// TIA Portal project "FS-DS-09" (V16) (continued)
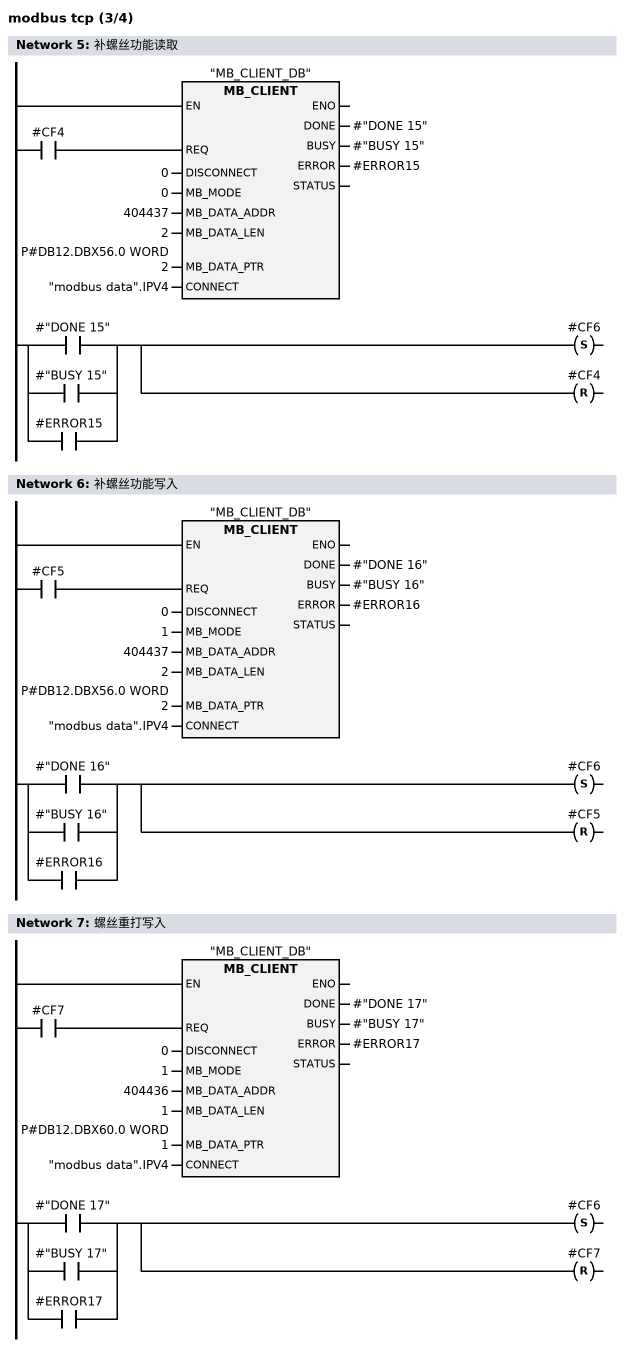
   "MB_CLIENT_DB"(REQ := #CF4,   // MB_CLIENT
                  DISCONNECT := 0,
                  MB_MODE := 0,
                  MB_DATA_ADDR := 404437,
                  MB_DATA_LEN := 2,
                  MB_DATA_PTR := P#DB12.DBX56.0 WORD 2,
                  CONNECT := "modbus data".IPV4,
                  DONE => #"DONE 15",
                  BUSY => #"BUSY 15",
                  ERROR => #ERROR15);
   IF #"DONE 15" OR #"BUSY 15" OR #ERROR15 THEN
       #CF6 := TRUE;
       #CF4 := FALSE;
   END_IF;
END_REGION

REGION Network 6: 补螺丝功能写入
   "MB_CLIENT_DB"(REQ := #CF5,   // MB_CLIENT
                  DISCONNECT := 0,
                  MB_MODE := 1,
                  MB_DATA_ADDR := 404437,
                  MB_DATA_LEN := 2,
                  MB_DATA_PTR := P#DB12.DBX56.0 WORD 2,
                  CONNECT := "modbus data".IPV4,
                  DONE => #"DONE 16",
                  BUSY => #"BUSY 16",
                  ERROR => #ERROR16);
   IF #"DONE 16" OR #"BUSY 16" OR #ERROR16 THEN
       #CF6 := TRUE;
       #CF5 := FALSE;
   END_IF;
END_REGION

REGION Network 7: 螺丝重打写入
   "MB_CLIENT_DB"(REQ := #CF7,   // MB_CLIENT
                  DISCONNECT := 0,
                  MB_MODE := 1,
                  MB_DATA_ADDR := 404436,
                  MB_DATA_LEN := 1,
                  MB_DATA_PTR := P#DB12.DBX60.0 WORD 1,
                  CONNECT := "modbus data".IPV4,
                  DONE => #"DONE 17",
                  BUSY => #"BUSY 17",
                  ERROR => #ERROR17);
   IF #"DONE 17" OR #"BUSY 17" OR #ERROR17 THEN
       #CF6 := TRUE;
       #CF7 := FALSE;
   END_IF;
END_REGION

REGION Network 8: 回原位标志位写入
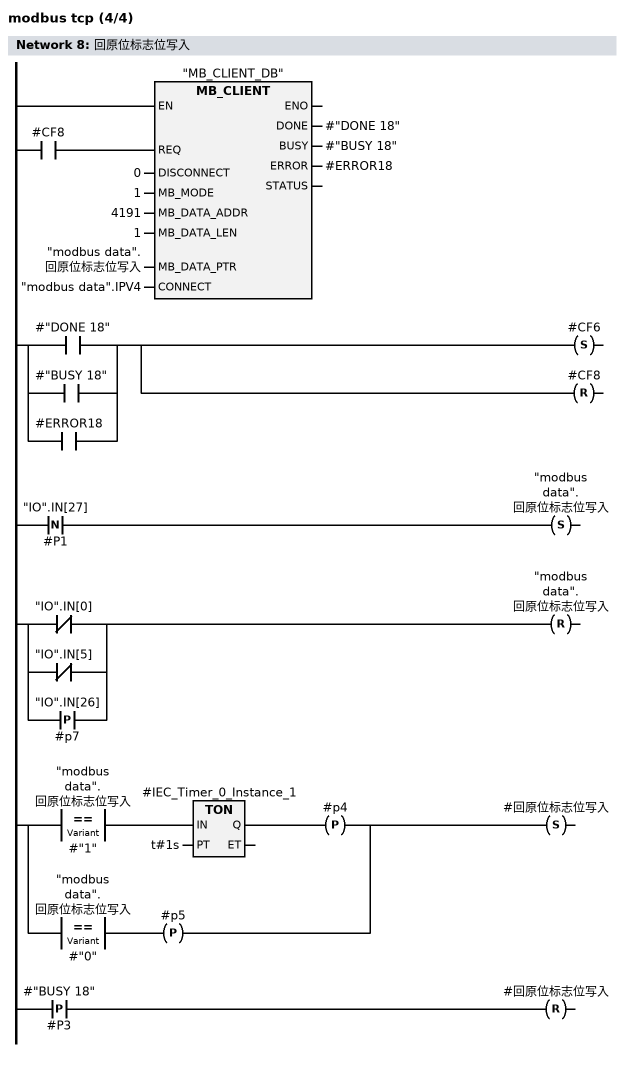
   "MB_CLIENT_DB"(REQ := #CF8,   // MB_CLIENT
                  DISCONNECT := 0,
                  MB_MODE := 1,
                  MB_DATA_ADDR := 4191,
                  MB_DATA_LEN := 1,
                  MB_DATA_PTR := "modbus data".回原位标志位写入,
                  CONNECT := "modbus data".IPV4,
                  DONE => #"DONE 18",
                  BUSY => #"BUSY 18",
                  ERROR => #ERROR18);
   IF #"DONE 18" OR #"BUSY 18" OR #ERROR18 THEN
       #CF6 := TRUE;
       #CF8 := FALSE;
   END_IF;
   #_w1 := NOT "IO".IN[27] AND #P1;   // falling edge of "IO".IN[27]
   #P1 := "IO".IN[27];
   IF #_w1 THEN "modbus data".回原位标志位写入 := TRUE; END_IF;
   #_w2 := "IO".IN[26] AND NOT #p7;   // rising edge of "IO".IN[26]
   #p7 := "IO".IN[26];
   IF NOT "IO".IN[0] OR NOT "IO".IN[5] OR #_w2 THEN "modbus data".回原位标志位写入 := FALSE; END_IF;
   #IEC_Timer_0_Instance_1(IN := "modbus data".回原位标志位写入 = #"1", PT := t#1s);   // TON
   #_w3 := #IEC_Timer_0_Instance_1.Q AND NOT #p4;   // rising edge
   #p4 := #IEC_Timer_0_Instance_1.Q;
   #_w4 := "modbus data".回原位标志位写入 = #"0";
   #_w5 := #_w4 AND NOT #p5;   // rising edge
   #p5 := #_w4;
   IF #_w3 OR #_w5 THEN #回原位标志位写入 := TRUE; END_IF;
   #_w6 := #"BUSY 18" AND NOT #P3;   // rising edge of #"BUSY 18"
   #P3 := #"BUSY 18";
   IF #_w6 THEN #回原位标志位写入 := FALSE; END_IF;
END_REGION

REGION Network 9 (SCL)
   "HengKongMC".hengkong.获取X轴当前坐标 := ("modbus data".Static_1.Static_1.X轴坐标/ 1000.0);
   "HengKongMC".hengkong.获取Y轴当前坐标 := "modbus data".Static_1.Static_1.Y轴坐标 / 1000.0;
   "HengKongMC".hengkong.获取Z轴当前坐标 := "modbus data".Static_1.Static_1.Z轴坐标 / 1000.0;
   "HengKongMC".hengkong.获取Y2轴当前坐标 := "modbus data".Static_1.Static_1.Y1轴坐标 / 1000.0;
   "HengKongMC".hengkong.螺丝孔加工完成情况查询 := "modbus data".Static_1.螺丝加工完成情况查询;
   "HengKongMC".hengkong.设备报警状态查询 := "modbus data".Static_1.设备报警状态查询;
   "HengKongMC".hengkong.左机加工完成情况查询 := "HengKongMC".hengkong.左机加工完成情况查询;
   "HengKongMC".hengkong.右机加工完成情况查询 := "modbus data".Static_1.右加工完成情况查询;
   "HengKongMC".hengkong.报警异常号 := WORD_TO_INT ("modbus data".Static_1.报警异常行号);
   IF "HMI".MU.HMI行号读取 OR "Control".MU.上位机行号读取 THEN
       "HengKongMC".hengkong.光标处运行标志 := WORD_TO_INT("modbus data".跳转行号.光标处运行标志);
       "HengKongMC".hengkong.当前程序所在行号 := WORD_TO_INT("modbus data".跳转行号.当前程序所在行号);
   END_IF;
   IF "HMI".MU.HMI行号写入 OR "Control".MU.上位机行号写入 THEN
       "modbus data".跳转行号.当前程序所在行号 := INT_TO_WORD("HengKongMC".hengkong.当前程序所在行号);
       "modbus data".跳转行号.光标处运行标志 := INT_TO_WORD("HengKongMC".hengkong.光标处运行标志);
   END_IF;
END_REGION
END_FUNCTION_BLOCK

// folder: 配方

FUNCTION_BLOCK "配方"   // FB6, LAD
{ S7_Optimized_Access := 'TRUE' }
VERSION : 0.1
BEGIN

REGION Network 1: 读
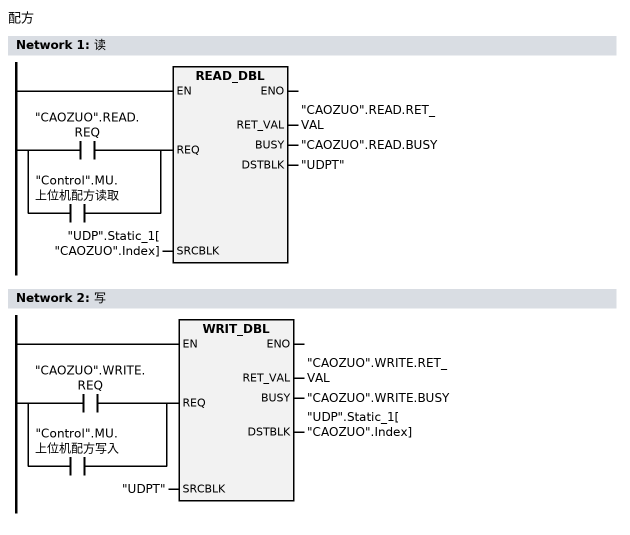
   "CAOZUO".READ.RET_VAL := READ_DBL(REQ := "CAOZUO".READ.REQ OR "Control".MU.上位机配方读取,
                           SRCBLK := "UDP".Static_1["CAOZUO".Index],
                           BUSY => "CAOZUO".READ.BUSY,
                           DSTBLK => "UDPT");
END_REGION

REGION Network 2: 写
   "CAOZUO".WRITE.RET_VAL := WRIT_DBL(REQ := "CAOZUO".WRITE.REQ OR "Control".MU.上位机配方写入,
                           SRCBLK := "UDPT",
                           BUSY => "CAOZUO".WRITE.BUSY,
                           DSTBLK => "UDP".Static_1["CAOZUO".Index]);
END_REGION

REGION Network 3 (SCL)
   IF "HMI".MU.HMI配方下载到PLC OR "Control".MU.上位机配方下载到PLC THEN
       "HMI".MU."PLC 配方名称" := "UDPT".加工文件名称;
       "HMI".MU."PLC 程序号" := "UDPT".加工文件编号;
       "HMI".MU.PLC螺丝个数 := "UDPT".加工螺丝数量;

   END_IF;
   IF NOT "IO".IN[4] AND  "吐钉模式".吐钉模式 AND NOT "HMI".工件完成信号 THEN
       "IO".OUT[6] := 1;
       "IO".OUT[7] := 1;
       "IO".OUT[8] :=1;
       "IO".OUT[9] := 1;
       "IO".OUT[10] := 1;
   ELSE
       "IO".OUT[6] := %DB10.DBX519.0;
       "IO".OUT[7] := %DB10.DBX519.1;
       "IO".OUT[8] := %DB10.DBX519.2;
       "IO".OUT[9] := %DB10.DBX519.3;
       "IO".OUT[10] := %DB10.DBX519.4;
   END_IF;
END_REGION
END_FUNCTION_BLOCK

(* ===== HMI "HMI_RT_1" =====
system functions are stored by id; their names below are inferred from use
connection "HMI_连接_1": ETHERNET, SMART_S7_1200_OMS

HMI tags "配方"
   "CAOZUO_READ_REQ" : Bool = PLC CAOZUO.READ.REQ AT %DB15.DBX0.0, 1 s
   "CAOZUO_WRITE_REQ" : Bool = PLC CAOZUO.WRITE.REQ AT %DB15.DBX6.0, 1 s
   "CAOZUO_Index" : Int = PLC CAOZUO.Index AT %DB15.DBW12, 1 s
   "UDPT_加工文件名称" : String[254] = PLC UDPT.加工文件名称 AT %DB14.DBX0.0, 1 s
   "HMI_MU_HMI配方下载到PLC" : Bool = PLC HMI.MU.HMI配方下载到PLC AT %DB10.DBX260.6, 1 s
   "HMI_MU_PLC 配方名称" : String[254] = PLC HMI.MU."PLC 配方名称" AT %DB10.DBX262.0, 1 s
   "HMI_MU_PLC 程序号" : Int = PLC HMI.MU."PLC 程序号" AT %DB10.DBW518, 1 s
   "UDPT_加工螺丝数量" : Int = PLC UDPT.加工螺丝数量 AT %DB14.DBW258, 1 s

HMI tags "输出"
   "三色灯黄色" : Bool = PLC IO.OUT[0] AT %DB1.DBX6.0, 1 s
   "三色灯绿色" : Bool = PLC IO.OUT[1] AT %DB1.DBX6.1, 1 s
   "三色灯红色" : Bool = PLC IO.OUT[2] AT %DB1.DBX6.2, 1 s
   "三色灯蜂鸣器" : Bool = PLC IO.OUT[3] AT %DB1.DBX6.3, 1 s
   "绿色半球指示灯" : Bool = PLC IO.OUT[4] AT %DB1.DBX6.4, 1 s
   "红色半球指示灯" : Bool = PLC IO.OUT[5] AT %DB1.DBX6.5, 1 s
   "运动控制卡任务选择1" : Bool = PLC IO.OUT[6] AT %DB1.DBX6.6, 1 s
   "运动控制卡任务选择2" : Bool = PLC IO.OUT[7] AT %DB1.DBX6.7, 1 s
   "运动控制卡任务选择3" : Bool = PLC IO.OUT[8] AT %DB1.DBX7.0, 1 s
   "运动控制卡任务选择4" : Bool = PLC IO.OUT[9] AT %DB1.DBX7.1, 1 s
   "运动控制卡任务选择5" : Bool = PLC IO.OUT[10] AT %DB1.DBX7.2, 1 s
   "Y1供料器有料输出" : Bool = PLC IO.OUT[11] AT %DB1.DBX7.3, 1 s
   "Y2供料器有料输出" : Bool = PLC IO.OUT[12] AT %DB1.DBX7.4, 1 s
   "运动控制卡启动" : Bool = PLC IO.OUT[13] AT %DB1.DBX7.5, 1 s
   "运动控制卡复位" : Bool = PLC IO.OUT[14] AT %DB1.DBX7.6, 1 s
   "运动控制卡紧急停止" : Bool = PLC IO.OUT[15] AT %DB1.DBX7.7, 1 s
   "运动控制卡停止" : Bool = PLC IO.OUT[16] AT %DB1.DBX8.0, 1 s
   "吸取螺丝电磁阀" : Bool = PLC IO.OUT[17] AT %DB1.DBX8.1, 1 s
   "下压气缸电磁阀" : Bool = PLC IO.OUT[18] AT %DB1.DBX8.2, 1 s
   "工装电磁铁" : Bool = PLC IO.OUT[19] AT %DB1.DBX8.3, 1 s
   "运动控制光栅报警" : Bool = PLC IO.OUT[20] AT %DB1.DBX8.4, 1 s
   "伺服复位" : Bool = PLC IO.OUT[21] AT %DB1.DBX8.5, 1 s
   "电批急停" : Bool = PLC IO.OUT[22] AT %DB1.DBX8.6, 1 s
   "备用(9)" : Bool = PLC IO.OUT[23] AT %DB1.DBX8.7, 1 s
   "FFU" : Bool = PLC IO.OUT[24] AT %DB1.DBX9.0, 1 s
   "照明" : Bool = PLC IO.OUT[25] AT %DB1.DBX9.1, 1 s
   "夹紧气缸1夹紧" : Bool = PLC IO.OUT[26] AT %DB1.DBX9.2, 1 s
   "夹紧气缸2夹紧" : Bool = PLC IO.OUT[27] AT %DB1.DBX9.3, 1 s
   "备用_3(1)" : Bool = PLC IO.OUT[28] AT %DB1.DBX9.4, 1 s
   "备用_4(1)" : Bool = PLC IO.OUT[29] AT %DB1.DBX9.5, 1 s
   "备用_5(1)" : Bool = PLC IO.OUT[30] AT %DB1.DBX9.6, 1 s
   "备用_6(1)" : Bool = PLC IO.OUT[31] AT %DB1.DBX9.7, 1 s
   "备用_7(1)" : Bool = PLC IO.OUT[32] AT %DB1.DBX10.0, 1 s
   "备用_8(1)" : Bool = PLC IO.OUT[33] AT %DB1.DBX10.1, 1 s

HMI tags "输入"
   "操作面板急停" : Bool = PLC IO.IN[0] AT %DB1.DBX0.0, 1 s
   "回原位" : Bool = PLC IO.IN[1] AT %DB1.DBX0.1, 1 s
   "启动按钮" : Bool = PLC IO.IN[2] AT %DB1.DBX0.2, 1 s
   "停止按钮" : Bool = PLC IO.IN[3] AT %DB1.DBX0.3, 1 s
   "手动/自动" : Bool = PLC IO.IN[4] AT %DB1.DBX0.4, 1 s
   "按钮盒急停" : Bool = PLC IO.IN[5] AT %DB1.DBX0.5, 1 s
   "左启动" : Bool = PLC IO.IN[6] AT %DB1.DBX0.6, 1 s
   "右启动" : Bool = PLC IO.IN[7] AT %DB1.DBX0.7, 1 s
   "安全门" : Bool = PLC IO.IN[8] AT %DB1.DBX1.0, 1 s
   "安全光幕" : Bool = PLC IO.IN[9] AT %DB1.DBX1.1, 1 s
   "Y1供料器有料" : Bool = PLC IO.IN[10] AT %DB1.DBX1.2, 1 s
   "Y2供料器有料" : Bool = PLC IO.IN[11] AT %DB1.DBX1.3, 1 s
   "1#工装产品信号" : Bool = PLC IO.IN[12] AT %DB1.DBX1.4, 1 s
   "2#工装产品信号" : Bool = PLC IO.IN[13] AT %DB1.DBX1.5, 1 s
   "气夹气缸到位2" : Bool = PLC IO.IN[14] AT %DB1.DBX1.6, 1 s
   "气夹气缸到位1" : Bool = PLC IO.IN[15] AT %DB1.DBX1.7, 1 s
   "工具错误" : Bool = PLC IO.IN[16] AT %DB1.DBX2.0, 1 s
   "工具拧紧OK" : Bool = PLC IO.IN[17] AT %DB1.DBX2.1, 1 s
   "工具拧紧NG" : Bool = PLC IO.IN[18] AT %DB1.DBX2.2, 1 s
   "工具准备好" : Bool = PLC IO.IN[19] AT %DB1.DBX2.3, 1 s
   "工具运行" : Bool = PLC IO.IN[20] AT %DB1.DBX2.4, 1 s
   "气源压力检测" : Bool = PLC IO.IN[21] AT %DB1.DBX2.5, 1 s
   "光栅屏蔽对射开关" : Bool = PLC IO.IN[22] AT %DB1.DBX2.6, 1 s
   "吸附信号" : Bool = PLC IO.IN[23] AT %DB1.DBX2.7, 1 s
   "电批下压气缸信号" : Bool = PLC IO.IN[24] AT %DB1.DBX3.0, 1 s
   "备用" : Bool = PLC IO.IN[25] AT %DB1.DBX3.1, 1 s
   "回原位中" : Bool = PLC IO.IN[26] AT %DB1.DBX3.2, 1 s
   "回原位完成" : Bool = PLC IO.IN[27] AT %DB1.DBX3.3, 1 s
   "X轴故障报警" : Bool = PLC IO.IN[28] AT %DB1.DBX3.4, 1 s
   "Y轴故障报警" : Bool = PLC IO.IN[29] AT %DB1.DBX3.5, 1 s
   "Z轴故障报警" : Bool = PLC IO.IN[30] AT %DB1.DBX3.6, 1 s
   "运动控制卡完成/释放夹紧气缸" : Bool = PLC IO.IN[31] AT %DB1.DBX3.7, 1 s
   "备用_3" : Bool = PLC IO.IN[32] AT %DB1.DBX4.0, 1 s
   "备用_4" : Bool = PLC IO.IN[33] AT %DB1.DBX4.1, 1 s
   "备用_5" : Bool = PLC IO.IN[34] AT %DB1.DBX4.2, 1 s
   "备用_6" : Bool = PLC IO.IN[35] AT %DB1.DBX4.3, 1 s
   "备用_7" : Bool = PLC IO.IN[36] AT %DB1.DBX4.4, 1 s
   "备用_8" : Bool = PLC IO.IN[37] AT %DB1.DBX4.5, 1 s
   "IO_IN{38}" : Bool = PLC IO.IN[38] AT %DB1.DBX4.6, 1 s
   "IO_IN{39}" : Bool = PLC IO.IN[39] AT %DB1.DBX4.7, 1 s
   "IO_IN{40}" : Bool = PLC IO.IN[40] AT %DB1.DBX5.0, 1 s

HMI tags "报警"
   "Alarm_运动控制板卡螺丝加工完成情况昂查询" : String[254] = PLC Alarm.运动控制板卡螺丝加工完成情况昂查询 AT %DB4.DBX0.0, 1 s
   "Alarm_运动控制板卡设备报警状态查询" : String[254] = PLC Alarm.运动控制板卡设备报警状态查询 AT %DB4.DBX256.0, 1 s
   "Alarm_运动控制板卡报警" : Bool = PLC Alarm.运动控制板卡报警 AT %DB4.DBX512.0, 1 s
   "Alarm_设备气源压力低报警" : Bool = PLC Alarm.设备气源压力低报警 AT %DB4.DBX512.1, 1 s
   "Alarm_面板急停报警" : Bool = PLC Alarm.面板急停报警 AT %DB4.DBX512.2, 1 s
   "Alarm_操作面板急停报警" : Bool = PLC Alarm.操作面板急停报警 AT %DB4.DBX512.3, 1 s
   "Alarm_安全门报警" : Bool = PLC Alarm.安全门报警 AT %DB4.DBX512.4, 1 s
   "Alarm_光幕报警" : Bool = PLC Alarm.光幕报警 AT %DB4.DBX512.5, 1 s
   "Alarm_回原位超时报警" : Bool = PLC Alarm.回原位超时报警 AT %DB4.DBX512.6, 1 s
   "Alarm_Y1供料器超时报警" : Bool = PLC Alarm.Y1供料器超时报警 AT %DB4.DBX512.7, 1 s
   "Alarm_Y2供料器超时报警" : Bool = PLC Alarm.Y2供料器超时报警 AT %DB4.DBX513.0, 1 s
   "Alarm_工装产品检测1无件报警" : Bool = PLC Alarm.工装产品检测1无件报警 AT %DB4.DBX513.1, 1 s
   "Alarm_工装产品检测2无件报警" : Bool = PLC Alarm.工装产品检测2无件报警 AT %DB4.DBX513.2, 1 s
   "Alarm_气缸夹紧1夹紧超时" : Bool = PLC Alarm.气缸夹紧1夹紧超时 AT %DB4.DBX513.3, 1 s
   "Alarm_气缸夹紧2夹紧超时" : Bool = PLC Alarm.气缸夹紧2夹紧超时 AT %DB4.DBX513.4, 1 s
   "Alarm_丹尼克尔错误报警" : Bool = PLC Alarm.丹尼克尔错误报警 AT %DB4.DBX513.5, 1 s
   "Alarm_一级报警" : Bool = PLC Alarm.一级报警 AT %DB4.DBX513.6, 1 s
   "Alarm_二级报警" : Bool = PLC Alarm.二级报警 AT %DB4.DBX513.7, 1 s
   "Alarm_下压气缸故障" : Bool = PLC Alarm.下压气缸故障 AT %DB4.DBX514.0, 1 s
   "Alarm_打螺丝延时过小" : Bool = PLC Alarm.打螺丝延时过小 AT %DB4.DBX514.1, 1 s
   "Alarm_真空检测失败" : Bool = PLC Alarm.真空检测失败 AT %DB4.DBX514.2, 1 s
   "Alarm_吸取螺丝失败" : Bool = PLC Alarm.吸取螺丝失败 AT %DB4.DBX514.3, 1 s
   "Alarm_分料超时" : Bool = PLC Alarm.分料超时 AT %DB4.DBX514.4, 1 s
   "Alarm_夹紧气缸故障FB运行前未复位" : Bool = PLC Alarm.夹紧气缸故障FB运行前未复位 AT %DB4.DBX514.5, 1 s
   "Alarm_下压气缸不在原位" : Bool = PLC Alarm.下压气缸不在原位 AT %DB4.DBX514.6, 1 s
   "Alarm_X轴故障报警" : Bool = PLC Alarm.X轴故障报警 AT %DB4.DBX514.7, 1 s
   "Alarm_Y轴故障报警" : Bool = PLC Alarm.Y轴故障报警 AT %DB4.DBX515.0, 1 s
   "Alarm_Z轴故障报警" : Bool = PLC Alarm.Z轴故障报警 AT %DB4.DBX515.1, 1 s

HMI tags "运动控制板卡"
   "HengKongMC_hengkong_DATA_获取X轴当前坐标" : LReal = PLC HengKongMC.hengkong.获取X轴当前坐标 AT %DB2.DBX6.0, 1 s
   "HengKongMC_hengkong_DATA_获取Y轴当前坐标" : LReal = PLC HengKongMC.hengkong.获取Y轴当前坐标 AT %DB2.DBX14.0, 1 s
   "HengKongMC_hengkong_DATA_获取Z轴当前坐标" : LReal = PLC HengKongMC.hengkong.获取Z轴当前坐标 AT %DB2.DBX22.0, 1 s
   "HengKongMC_hengkong_报警异常号" : Int = PLC HengKongMC.hengkong.报警异常号 AT %DB2.DBW52, 1 s
   "HengKongMC_hengkong_光标处运行标志" : Int = PLC HengKongMC.hengkong.光标处运行标志 AT %DB2.DBW54, 1 s
   "HengKongMC_hengkong_当前程序所在行号" : Int = PLC HengKongMC.hengkong.当前程序所在行号 AT %DB2.DBW56, 1 s
   "HengKongMC_hengkong_补螺丝功能_读取" : Bool = PLC HMI.MU.HMI行号读取 AT %DB10.DBX260.4, 1 s
   "HengKongMC_hengkong_补螺丝功能_写入" : Bool = PLC HMI.MU.HMI行号写入 AT %DB10.DBX260.3, 1 s

HMI tags "HMI控制"
   "HMI_MU_HMI吸附电磁阀" : Bool = PLC HMI.MU.HMI吸附电磁阀 AT %DB10.DBX0.0, 1 s
   "HMI_MU_HMI下压气缸电磁阀" : Bool = PLC HMI.MU.HMI下压气缸电磁阀 AT %DB10.DBX0.1, 1 s
   "HMI_MU_HMI停止" : Bool = PLC HMI.MU.HMI停止 AT %DB10.DBX0.2, 1 s
   "HMI_MU_HMIFFU" : Bool = PLC HMI.MU.HMIFFU AT %DB10.DBX0.3, 1 s
   "HMI_MU_HMI照明" : Bool = PLC HMI.MU.HMI照明 AT %DB10.DBX0.4, 1 s
   "HMI_MU_HMI夹紧气缸1夹紧" : Bool = PLC HMI.MU.HMI夹紧气缸1夹紧 AT %DB10.DBX0.5, 1 s
   "HMI_MU_HMI夹紧气缸2夹紧" : Bool = PLC HMI.MU.HMI夹紧气缸2夹紧 AT %DB10.DBX0.6, 1 s
   "HMI_MU_HMI机消音" : Bool = PLC HMI.MU.HMI机消音 AT %DB10.DBX0.7, 1 s
   "HMI_MU_HMI伺服错误复位" : Bool = PLC HMI.MU.HMI伺服错误复位 AT %DB10.DBX1.0, 1 s
   "HMI_MU_HMI加工文件选择" : Int = PLC HMI.MU.HMI加工文件选择 AT %DB10.DBW2, 1 s
   "HMI_MU_HMI加工文件名称" : String[254] = PLC HMI.MU.HMI加工文件名称 AT %DB10.DBX4.0, 1 s
   "HMI_MU_HMI启动信号" : Bool = PLC HMI.MU.HMI启动信号 AT %DB10.DBX260.0, 1 s
   "HMI_MU_MHI屏蔽信号" : Bool = PLC HMI.MU.MHI屏蔽信号 AT %DB10.DBX260.1, 1 s
   "HMI_MU_HMI电批启动" : Bool = PLC HMI.MU.HMI电批启动 AT %DB10.DBX260.2, 1 s
   "HMI_MU_HMI行号写入" : Bool = PLC HMI.MU.HMI行号写入 AT %DB10.DBX260.3, 1 s
   "HMI_MU_HMI行号读取" : Bool = PLC HMI.MU.HMI行号读取 AT %DB10.DBX260.4, 1 s
   "HMI_MU_HMI工装电磁铁启动" : Bool = PLC HMI.MU.HMI工装电磁铁启动 AT %DB10.DBX260.5, 1 s
   "HMI_MU_HMI计数器清零" : Bool = PLC HMI.MU.HMI计数器清零 AT %DB10.DBX522.0, 1 s
   "HMI_MU_HMI合格" : Real = PLC HMI.MU.HMI合格 AT %DB10.DBD524, 1 s
   "HMI_MU_HMI 不合格" : Real = PLC HMI.MU."HMI 不合格" AT %DB10.DBD528, 1 s
   "HMI_MU_HMI合格率" : Real = PLC HMI.MU.HMI合格率 AT %DB10.DBD532, 1 s
   "HMI_MU_HMI 产品数" : Real = PLC HMI.MU."HMI 产品数" AT %DB10.DBD536, 1 s
   "HMI_MU_HMI 运行螺丝个数" : Int = PLC HMI.MU."HMI 运行螺丝个数" AT %DB10.DBW540, 1 s
   "HMI_HMI 运行螺丝个数NG" : Int = PLC HMI."HMI 运行螺丝个数NG" AT %DB10.DBW544, 1 s
   "HMI_工件完成信号" : Bool = PLC HMI.工件完成信号 AT %DB10.DBX546.0, 1 s
   "吐钉模式_吐钉模式" : Bool = PLC 吐钉模式.吐钉模式 AT %DB1.DBX0.0, 1 s

HMI tags "hmi 报警"
   "HMI_Tag_1" : Word AT %DB4.DBW512, 500 ms
   "HMI_Tag_2" : Word AT %DB4.DBW514, 500 ms
   "HMI_Tag_3" : Word AT %DB4.DBW516, 500 ms
   "HMI_Tag_4" : Word AT %DB7.DBW0, 1 s

HMI tags "内部变量"
   "跳转画面" : Int, internal
   "屏蔽菜单" : Int, internal
   "报警消除" : Int, internal
   "隐藏画面" : Int, internal

HMI tags "运动控制板卡输入IO"
   "HengKongMC_输入_X轴原位" : Bool = PLC HengKongMC.输入.X轴原位 AT %DB2.DBX0.0, 1 s
   "HengKongMC_输入_Y轴原位" : Bool = PLC HengKongMC.输入.Y轴原位 AT %DB2.DBX0.1, 1 s
   "HengKongMC_输入_Z轴原位" : Bool = PLC HengKongMC.输入.Z轴原位 AT %DB2.DBX0.2, 1 s
   "HengKongMC_输入_X4备用" : Bool = PLC HengKongMC.输入.X4备用 AT %DB2.DBX0.3, 1 s
   "HengKongMC_输入_Y2供料器有料" : Bool = PLC HengKongMC.输入.Y2供料器有料 AT %DB2.DBX0.4, 1 s
   "HengKongMC_输入_电批启动" : Bool = PLC HengKongMC.输入.电批启动 AT %DB2.DBX0.5, 1 s
   "HengKongMC_输入_任务选择1" : Bool = PLC HengKongMC.输入.任务选择1 AT %DB2.DBX0.6, 1 s
   "HengKongMC_输入_任务选择2" : Bool = PLC HengKongMC.输入.任务选择2 AT %DB2.DBX0.7, 1 s
   "HengKongMC_输入_启动" : Bool = PLC HengKongMC.输入.启动 AT %DB2.DBX1.0, 1 s
   "HengKongMC_输入_回原位" : Bool = PLC HengKongMC.输入.回原位 AT %DB2.DBX1.1, 1 s
   "HengKongMC_输入_急停" : Bool = PLC HengKongMC.输入.急停 AT %DB2.DBX1.2, 1 s
   "HengKongMC_输入_OK" : Bool = PLC HengKongMC.输入.OK AT %DB2.DBX1.3, 1 s
   "HengKongMC_输入_光幕和门控报警" : Bool = PLC HengKongMC.输入.光幕和门控报警 AT %DB2.DBX1.4, 1 s
   "HengKongMC_输入_任务选择3" : Bool = PLC HengKongMC.输入.任务选择3 AT %DB2.DBX1.5, 1 s
   "HengKongMC_输入_任务选择4" : Bool = PLC HengKongMC.输入.任务选择4 AT %DB2.DBX1.6, 1 s
   "HengKongMC_输入_任务选择5" : Bool = PLC HengKongMC.输入.任务选择5 AT %DB2.DBX1.7, 1 s
   "HengKongMC_输入_负压传感器" : Bool = PLC HengKongMC.输入.负压传感器 AT %DB2.DBX2.0, 1 s
   "HengKongMC_输入_Y1供料器有料" : Bool = PLC HengKongMC.输入.Y1供料器有料 AT %DB2.DBX2.1, 1 s
   "HengKongMC_输入_X19" : Bool = PLC HengKongMC.输入.X19 AT %DB2.DBX2.2, 1 s
   "HengKongMC_输入_X20" : Bool = PLC HengKongMC.输入.X20 AT %DB2.DBX2.3, 1 s
   "HengKongMC_输入_X21" : Bool = PLC HengKongMC.输入.X21 AT %DB2.DBX2.4, 1 s
   "HengKongMC_输入_下压气缸原位" : Bool = PLC HengKongMC.输入.下压气缸原位 AT %DB2.DBX2.5, 1 s
   "HengKongMC_输入_X23" : Bool = PLC HengKongMC.输入.X23 AT %DB2.DBX2.6, 1 s
   "HengKongMC_输入_停止" : Bool = PLC HengKongMC.输入.停止 AT %DB2.DBX2.7, 1 s

HMI tags "运动控制板卡输出IO"
   "HengKongMC_输出_吸取螺丝信号" : Bool = PLC HengKongMC.输出.吸取螺丝信号 AT %DB2.DBX4.0, 1 s
   "HengKongMC_输出_回原位成功" : Bool = PLC HengKongMC.输出.回原位成功 AT %DB2.DBX4.1, 1 s
   "HengKongMC_输出_回原位中" : Bool = PLC HengKongMC.输出.回原位中 AT %DB2.DBX4.2, 1 s
   "HengKongMC_输出_下压气缸信号" : Bool = PLC HengKongMC.输出.下压气缸信号 AT %DB2.DBX4.3, 1 s
   "HengKongMC_输出_Y5" : Bool = PLC HengKongMC.输出.Y5 AT %DB2.DBX4.4, 1 s
   "HengKongMC_输出_认螺帽反转" : Bool = PLC HengKongMC.输出.认螺帽反转 AT %DB2.DBX4.5, 1 s
   "HengKongMC_输出_Y7" : Bool = PLC HengKongMC.输出.运动控制卡完成信号 AT %DB2.DBX4.6, 1 s
   "HengKongMC_输出_Y8" : Bool = PLC HengKongMC.输出.Y8 AT %DB2.DBX4.7, 1 s
   "HengKongMC_输出_任务选择0" : Bool = PLC HengKongMC.输出.任务选择0 AT %DB2.DBX5.0, 1 s
   "HengKongMC_输出_任务选择1" : Bool = PLC HengKongMC.输出.任务选择1 AT %DB2.DBX5.1, 1 s
   "HengKongMC_输出_任务选择2" : Bool = PLC HengKongMC.输出.任务选择2 AT %DB2.DBX5.2, 1 s
   "HengKongMC_输出_Y12" : Bool = PLC HengKongMC.输出.Y12 AT %DB2.DBX5.3, 1 s
   "HengKongMC_输出_启动电批" : Bool = PLC HengKongMC.输出.启动电批 AT %DB2.DBX5.4, 1 s
   "HengKongMC_输出_Y14" : Bool = PLC HengKongMC.输出.Y14 AT %DB2.DBX5.5, 1 s
   "回原位标志位" : Bool = PLC HengKongMC.输出.回原位标志位 AT %DB2.DBX5.6, 1 s
   "HengKongMC_输出_Y16" : Bool = PLC HengKongMC.输出.Y16 AT %DB2.DBX5.7, 1 s

HMI tags "屏蔽"
   "Blocking function_Y1供料器报警屏蔽" : Bool = PLC "Blocking function".Y1供料器报警屏蔽 AT %DB7.DBX0.0, 1 s
   "Blocking function_Y2供料器报警屏蔽" : Bool = PLC "Blocking function".Y2供料器报警屏蔽 AT %DB7.DBX0.1, 1 s
   "Blocking function_工装产品检测1屏蔽" : Bool = PLC "Blocking function".工装产品检测1屏蔽 AT %DB7.DBX0.2, 1 s
   "Blocking function_工装产品检测2屏蔽" : Bool = PLC "Blocking function".工装产品检测2屏蔽 AT %DB7.DBX0.3, 1 s
   "Blocking function_夹紧气缸1夹紧屏蔽" : Bool = PLC "Blocking function".夹紧气缸1夹紧屏蔽 AT %DB7.DBX0.4, 1 s
   "Blocking function_夹紧气缸2夹紧屏蔽" : Bool = PLC "Blocking function".夹紧气缸2夹紧屏蔽 AT %DB7.DBX0.5, 1 s
   "Blocking function_上位机屏蔽" : Bool = PLC "Blocking function".上位机屏蔽 AT %DB7.DBX0.6, 1 s
   "Blocking function_安全门屏蔽" : Bool = PLC "Blocking function".安全门屏蔽 AT %DB7.DBX0.7, 1 s
   "Blocking function_光幕屏蔽" : Bool = PLC "Blocking function".光幕屏蔽 AT %DB7.DBX1.0, 1 s

HMI tags "伺服状态"
   "负方向x" : Bool = PLC 负方向x AT %I6.2, 1 s
   "正方向x" : Bool = PLC 正方向x AT %I6.3, 1 s
   "准备OKx" : Bool = PLC 准备OKx AT %I42.0, 1 s
   "故障报警x" : Bool = PLC 故障报警x AT %I42.1, 1 s
   "故障代码x" : DWord = PLC 故障代码x AT %ID17, 1 s
   "负方向y" : Bool = PLC 负方向y AT %I10.2, 1 s
   "正方向y" : Bool = PLC 正方向y AT %I10.3, 1 s
   "准备OKy" : Bool = PLC 准备OKy AT %I46.0, 1 s
   "故障报警y" : Bool = PLC 故障报警y AT %I46.1, 1 s
   "故障代码y" : DWord = PLC 故障代码y AT %ID21, 1 s
   "负方向z" : Bool = PLC 负方向z AT %I14.2, 1 s
   "正方向z" : Bool = PLC 正方向z AT %I14.3, 1 s
   "准备OKz" : Bool = PLC 准备OKz AT %I50.0, 1 s
   "故障报警z" : Bool = PLC 故障报警z AT %I50.1, 1 s
   "故障代码z" : DWord = PLC 故障代码z AT %ID25, 1 s

HMI tags "系统时间"
   "系统时间_SET" : Bool = PLC 系统时间.SET, 1 s
   "系统时间_WRDT" : DTL = PLC 系统时间.WRDT, 1 s
   "系统时间_RDDT" : DTL = PLC 系统时间.RDDT, 1 s
   "系统时间_RET1" : Word = PLC 系统时间.RET1, 1 s
   "系统时间_RET2" : Word = PLC 系统时间.RET2, 1 s

discrete alarms
   2: '设备气源压力低报警', class Errors, trigger "HMI_Tag_1" bit 9
   3: '面板急停报警', class Errors, trigger "HMI_Tag_1" bit 10
   4: '操作面板急停报警', class Errors, trigger "HMI_Tag_1" bit 11
   5: '安全门报警', class Errors, trigger "HMI_Tag_1" bit 12
   6: '光幕报警', class Errors, trigger "HMI_Tag_1" bit 13
   7: '回原位超时报警', class Errors, trigger "HMI_Tag_1" bit 14
   8: 'Y1供料器超时报警', class Errors, trigger "HMI_Tag_1" bit 15
   9: 'Y2供料器超时报警', class Errors, trigger "HMI_Tag_1" bit 0
   10: '工装产品检测1无件报警', class Errors, trigger "HMI_Tag_1" bit 1
   11: '工装产品检测2无件报警', class Errors, trigger "HMI_Tag_1" bit 2
   12: '气缸夹紧1夹紧超时', class Errors, trigger "HMI_Tag_1" bit 3
   13: '气缸夹紧2夹紧超时', class Errors, trigger "HMI_Tag_1" bit 4
   14: '丹尼克尔错误报警', class Errors, trigger "HMI_Tag_1" bit 5
   15: '一级报警', class Errors, trigger "HMI_Tag_1" bit 6
   16: '二级报警', class Errors, trigger "HMI_Tag_1" bit 7
   17: '下压气缸故障', class Errors, trigger "HMI_Tag_2" bit 8
   18: '打螺丝延时过小', class Errors, trigger "HMI_Tag_2" bit 9
   19: '真空检测失败', class Errors, trigger "HMI_Tag_2" bit 10
   20: '吸取螺丝失败', class Errors, trigger "HMI_Tag_2" bit 11
   21: '分料超时', class Errors, trigger "HMI_Tag_2" bit 12
   22: '夹紧气缸故障FB运行前未复位', class Errors, trigger "HMI_Tag_2" bit 13
   23: '下压气缸不在原位', class Errors, trigger "HMI_Tag_2" bit 14
   24: 'X轴故障报警', class Errors, trigger "HMI_Tag_2" bit 15
   25: 'Y轴故障报警', class Errors, trigger "HMI_Tag_2" bit 0
   26: 'Z轴故障报警', class Errors, trigger "HMI_Tag_2" bit 1
   27: 'Y1供料器报警屏蔽开启', class Warnings, trigger "HMI_Tag_4" bit 8
   28: 'Y2供料器报警屏蔽开启', class Warnings, trigger "HMI_Tag_4" bit 9
   29: '工装产品检测1屏蔽开启', class Warnings, trigger "HMI_Tag_4" bit 10
   30: '工装产品检测2屏蔽开启', class Warnings, trigger "HMI_Tag_4" bit 11
   31: '夹紧气缸1夹紧屏蔽开启', class Warnings, trigger "HMI_Tag_4" bit 12
   32: '夹紧气缸2夹紧屏蔽开启', class Warnings, trigger "HMI_Tag_4" bit 13
   33: '上位机屏蔽开启', class Warnings, trigger "HMI_Tag_4" bit 14
   34: '安全门屏蔽开启', class Warnings, trigger "HMI_Tag_4" bit 15
   35: '光幕屏蔽开启', class Warnings, trigger "HMI_Tag_4" bit 0

text list "产品切换": 0 'Part_0'; 1 'Part_1'; 2 'Part_2'; 3 'Part_3'; 4 'Part_4'; 5 'Part_5'; 6 'Part_6'; 7 'Part_7'; 8 'Part_8'; 9 'Part_9'; 10 'Part_10'; 11 'Part_11'; 12 'Part_12'; 13 'Part_13'; 14 'Part_14'; 15 'Part_15'; 16 'Part_16'; 17 'Part_17'; 18 'Part_18'; 19 'Part_19'; 20 'Part_20'; 21 'Part_21'; 22 'Part_22'; 23 'Part_23'; 24 'Part_24'; 25 'Part_25'; 26 'Part_26'; 27 'Part_27'; 28 'Part_28'; 29 'Part_29'; 30 'Part_30'

text list "product_list": 1 'AT005'; 2 'Part_2'; 3 'Part_3'; 4 'Part_4'; 5 'Part_5'; 6 'Part_6'; 7 'Part_7'; 8 'Part_8'; 9 'Part_9'; 10 'Part_10'; 11 'Part_11'; 12 'Part_12'; 13 'Part_13'

text list "信号监控": 12 'I0.0-I1.5'; 13 'I2.0-I2.7'; 14 'I3.0-I3.7'; 15 'I4.0-I4.7'; 16 'Q0.0-Q1.1'; 17 'Q2.0-Q2.7'; 18 'Q3.0-Q3.7'; 19 'Q4.0-Q4.7'; 20 '板卡X1-X15'; 21 '板卡X16-X24'; 22 '板卡Y1-Y15'; 23 '板卡Y16'; 24 ''

text list "屏蔽信号": 0 '取消屏蔽'; 1 '开启屏蔽'

text list "屏蔽菜单": 2 '菜单一'; 26 '菜单二'

text list "加工螺丝": 0 ''; 1 '第1个螺丝完成'; 2 '第2个螺丝完成'; 3 '第3个螺丝完成'; 4 '第4个螺丝完成'; 5 '第5个螺丝完成'; 6 '第6个螺丝完成'; 7 '第7个螺丝完成'; 8 '第8个螺丝完成'; 9 '第9个螺丝完成'; 10 '第10个螺丝完成'; 11 '第11个螺丝完成'; 12 '第12个螺丝完成'; 13 '第13个螺丝完成'; 14 '第14个螺丝完成'; 15 '第15个螺丝完成'; 16 '第16个螺丝完成'; 17 '第17个螺丝完成'; 18 '第18个螺丝完成'; 19 '第19个螺丝完成'; 20 '第20个螺丝完成'; 21 '第21个螺丝完成'; 22 '第22个螺丝完成'; 23 '第23个螺丝完成'; 24 '第24个螺丝完成'; 25 '第25个螺丝完成'; 26 '第26个螺丝完成'; 27 '第27个螺丝完成'; 28 '第28个螺丝完成'; 29 '第29个螺丝完成'; 30 '第30个螺丝完成'

text list "加工螺丝_1": 0 ''; 1 '第1个螺丝NG'; 2 '第2个螺丝NG'; 3 '第3个螺丝NG'; 4 '第4个螺丝NG'; 5 '第5个螺丝NG'; 6 '第6个螺丝NG'; 7 '第7个螺丝NG'; 8 '第8个螺丝NG'; 9 '第9个螺丝NG'; 10 '第10个螺丝NG'; 11 '第11个螺丝NG'; 12 '第12个螺丝NG'; 13 '第13个螺丝NG'; 14 '第14个螺丝NG'; 15 '第15个螺丝NG'; 16 '第16个螺丝NG'; 17 '第17个螺丝NG'; 18 '第18个螺丝NG'; 19 '第19个螺丝NG'; 20 '第20个螺丝NG'; 21 '第21个螺丝NG'; 22 '第22个螺丝NG'; 23 '第23个螺丝NG'; 24 '第24个螺丝NG'; 25 '第25个螺丝NG'; 26 '第26个螺丝NG'; 27 '第27个螺丝NG'; 28 '第28个螺丝NG'; 29 '第29个螺丝NG'; 30 '第30个螺丝NG'

screen "主页" 800x480, template "按钮"
   GraphicView "图形视图_2" at 159,66 size 50x50; Picture "图形_2"
   Rectangle "模板_矩形_5" at 586,219 size 170x100
      Visibility <- "HMI_工件完成信号"
   TextField "文本域_1" at 654,254 size 33x29; Text 'OK'
      Visibility <- "HMI_工件完成信号"
   TextField "文本域_7" at 219,187 size 93x35; Text '产品SN码'
   IOField "I/O 域_4" at 220,227 size 312x35; FormatPattern ?????????????????????????
   TextField "文本域_6" at 219,281 size 85x23; Text '产品选择'
   SymbolicIOField "符号 I/O 域_1" at 220,305 size 160x35; TextOn '1'; TextOff '0'; TextList "产品切换"
      ProcessValue <- "CAOZUO_Index"
   Button "HmiScreenItemData_12" at 395,366 size 127x35; TextOff '下载PLC'; PictureOn "图形_13"; PictureOff "图形_38"
      on Press: SetBit("HMI_MU_HMI配方下载到PLC")
      on Release: ResetBit("HMI_MU_HMI配方下载到PLC")
      Visibility <- "手动/自动"
   IOField "I/O 域_5" at 220,366 size 160x35; FormatPattern ??????????
      ProcessValue <- "UDPT_加工文件名称"
   TextField "文本域_10" at 219,341 size 85x23; Text '产品名称'
   Rectangle "模板_矩形_1" at 586,219 size 170x100
      Visibility <- "HMI_工件完成信号"
   TextField "文本域_9" at 654,254 size 33x29; Text 'OK'
      Visibility <- "HMI_工件完成信号"
   Button "HmiScreenItemData_1" at 394,305 size 127x35; TextOff '读取'; PictureOff "图形_38"; PictureOn "图形_13"
      on Press: SetBit("CAOZUO_READ_REQ")
      on Release: ResetBit("CAOZUO_READ_REQ")
      Visibility <- "手动/自动"
   Button "模板_按钮_2" at 221,138 size 96x32; TextOn '计数清零'; TextOff '计数清零'; Authorization "User"
      on Press: SetBit("HMI_MU_HMI计数器清零")
      on Release: ResetBit("HMI_MU_HMI计数器清零")
      Visibility <- "隐藏画面"
   Button "模板_按钮_3" at 423,137 size 96x32; TextOn '取消'; TextOff '取消'
      Visibility <- "隐藏画面"
      on Press: SetTag("隐藏画面", 0)
   TextField "模板_文本域_1" at 220,76 size 73x20; Text '产品计数'
   TextField "模板_文本域_2" at 297,76 size 57x20; Text 'OK计数'
   TextField "模板_文本域_3" at 372,76 size 57x20; Text 'NG计数'
   TextField "模板_文本域_4" at 445,76 size 56x20; Text '合格率'
   IOField "模板_I/O 域_4" at 220,101 size 71x23; FormatPattern s99999
      ProcessValue <- "HMI_MU_HMI 产品数"
   IOField "模板_I/O 域_6" at 295,101 size 71x23; FormatPattern s99999
      ProcessValue <- "HMI_MU_HMI合格"
   IOField "模板_I/O 域_7" at 368,101 size 71x23; FormatPattern s99999
      ProcessValue <- "HMI_MU_HMI 不合格"
   IOField "模板_I/O 域_8" at 443,101 size 71x23; FormatPattern s999.9; Unit %
      ProcessValue <- "HMI_MU_HMI合格率"
   Button "模板_按钮_1" at 216,67 size 306x68; TextOff 'Text'
      on Press: SetTag("隐藏画面", 1)
   IOField "I/O 域_6" at 219,427 size 160x35; FormatPattern s99
      ProcessValue <- "UDPT_加工螺丝数量"
   TextField "文本域_8" at 219,402 size 105x23; Text '锁螺丝个数'
   TextField "文本域_12" at 556,429 size 230x40; Text '* 按停止按钮后回原位或取 下当前螺丝后按启动键重打。'
      Visibility <- "红色半球指示灯"
   Group "Group" at 586,322 size 170x100
   Group "Group_1" at 586,322 size 170x100
   SymbolicIOField "符号 I/O 域_2" at 586,148 size 160x35; TextOff '0'; TextOn '1'; TextList "加工螺丝"
      ProcessValue <- "HMI_MU_HMI 运行螺丝个数"
   TextField "文本域_3" at 586,118 size 133x35; Text '螺丝加工状态'
   TextField "文本域_4" at 586,55 size 133x35; Text '螺丝加工数量'
   IOField "I/O 域_1" at 586,84 size 160x35; FormatPattern 99
      ProcessValue <- "UDPT_加工螺丝数量"
   SymbolicIOField "符号 I/O 域_3" at 586,181 size 160x35; TextOn '1'; TextOff '0'; TextList "加工螺丝_1"
      ProcessValue <- "HMI_HMI 运行螺丝个数NG"
   Button "HmiScreenItemData_2" at 395,427 size 127x35; TextOff '吐钉'; PictureOn "图形_13"; PictureOff "图形_38"
      on Press: SetBit("吐钉模式_吐钉模式")
      Visibility <- "手动/自动"
      Appearance <- "吐钉模式_吐钉模式"
   Rectangle "模板_矩形_6" at 586,322 size 170x100
      Visibility <- "红色半球指示灯"
   TextField "文本域_2" at 654,357 size 33x29; Text 'NG'
      Visibility <- "红色半球指示灯"
   Rectangle "模板_矩形_2" at 586,322 size 170x100
      Visibility <- "红色半球指示灯"
   TextField "文本域_11" at 654,357 size 33x29; Text 'NG'
      Visibility <- "红色半球指示灯"

Template "按钮" 800x480
   GraphicView "模板_图形视图_1" at 0,0 size 102x59; Picture "33"
   GraphicView "模板_图形视图_3" at 102,0 size 697x59; Picture "33"
   Group "Group" at 0,0 size 799x59; Picture "LOGO"
   GraphicView "模板_图形视图_2" at 0,0 size 200x59; Picture "复赛"
   Button "HmiScreenItemData_1" at 11,68 size 143x47; TextOn '主页'; TextOff '主页'; PictureOff "图形_12"; PictureOn "图形_12"
      on Release: ActivateScreen("主页", 0)
   Button "HmiScreenItemData_2" at 11,187 size 143x47; TextOn '手动控制'; TextOff '手动控制'; PictureOn "图形_9"; PictureOff "图形_9"; Authorization "User"
      on Release: ActivateScreen("气缸控制", 0)
   Button "HmiScreenItemData_3" at 11,307 size 143x47; TextOff '屏蔽管理'; PictureOff "图形_23"; PictureOn "图形_23"; Authorization "User"
      on Release: ActivateScreen("屏蔽管理", 0)
   Button "HmiScreenItemData_5" at 11,127 size 143x47; TextOn '信号监控'; TextOff '信号监控'; PictureOn "Navigates to SIMATIC PLC 监视表 for TP700 Comfort 14.0.1.0"; PictureOff "Navigates to SIMATIC PLC 监视表 for TP700 Comfort 14.0.1.0"
      on Release: ActivateScreen("信号监控", 0)
   Button "HmiScreenItemData_8" at 11,427 size 143x47; TextOn '下一页'; TextOff '下一页'; PictureOff "图形_15"; PictureOn "图形_15"
      on Release: ActivateScreen("主页_1", 0)
   Button "HmiScreenItemData_11" at 11,247 size 143x47; TextOff '产品管理'; PictureOff "Navigates to 项目信息 for TP700 Comfort 14.0.1.0"; PictureOn "Navigates to 项目信息 for TP700 Comfort 14.0.1.0"; Authorization "User"
      on Release: ActivateScreen("配方", 0)
   Button "HmiScreenItemData_7" at 11,367 size 143x47; TextOn '伺服状态'; TextOff '伺服状态'; PictureOff "图形_10"; PictureOn "图形_10"
      on Release: ActivateScreen("伺服状态", 0)
   IOField "模板_I/O 域_1" at 258,13 size 85x32; FormatPattern ????????????????????????????????????????????????????????????????????????????????
      ProcessValue <- "HMI_MU_PLC 配方名称"
   IOField "模板_I/O 域_2" at 362,15 size 35x30; FormatPattern 99
      ProcessValue <- "HMI_MU_PLC 程序号"
   TextField "文本域_6" at 410,16 size 91x29; Text '回原位中'
      Visibility <- "回原位中"
   TextField "文本域_2" at 501,16 size 91x29; Text '请回原位'
      Visibility <- "回原位标志位"
      Appearance <- "回原位标志位"
   TextField "文本域_1" at 410,16 size 111x29; Text '回原位完成'
      Visibility <- "回原位标志位"
   DateTimeField "模板_日期/时间域_1" at 597,20 size 201x21

screen "气缸控制" 800x480, template "按钮"
   TextField "文本域_1" at 259,76 size 39x20; Text '状态'
   TextField "文本域_2" at 421,76 size 73x20; Text '注释名称'
   TextField "文本域_3" at 639,76 size 73x20; Text '操作按钮'
   Group "Group" at 211,67 size 571x402
   Switch "开关_5" at 622,374 size 100x40; TextOn '开启'; CaptionText 'Switch'; TextOff '开启'
      ProcessValue <- "HMI_MU_HMIFFU"
      Appearance <- "FFU"
   GraphicView "图形视图_2" at 159,185 size 50x50; Picture "图形_2"
   Switch "开关_1" at 622,111 size 100x40; CaptionText 'Switch'; TextOff '开启'; TextOn '开启'
      ProcessValue <- "HMI_MU_HMI夹紧气缸1夹紧"
      Visibility <- "手动/自动"
      Appearance <- "备用_3(1)"
   Switch "开关_3" at 622,270 size 100x40; TextOn '开启'; CaptionText 'Switch'; TextOff '开启'
      ProcessValue <- "HMI_MU_HMI下压气缸电磁阀"
      Appearance <- "下压气缸电磁阀"
      Visibility <- "手动/自动"
   Switch "开关_4" at 622,217 size 100x40; TextOn '开启'; CaptionText 'Switch'; TextOff '开启'
      ProcessValue <- "HMI_MU_HMI吸附电磁阀"
      Appearance <- "吸取螺丝电磁阀"
      Visibility <- "手动/自动"
   Switch "开关_6" at 622,428 size 100x40; TextOn '开启'; CaptionText 'Switch'; TextOff '开启'
      ProcessValue <- "HMI_MU_HMI照明"
      Appearance <- "照明"
   Switch "开关_7" at 622,164 size 100x40; TextOn '开启'; CaptionText 'Switch'; TextOff '开启'
      Appearance <- "工装电磁铁"
      ProcessValue <- "HMI_MU_HMI工装电磁铁启动"
      Visibility <- "手动/自动"
   TextField "文本域_6" at 410,122 size 85x23; Text '工装夹紧'
   TextField "文本域_4" at 410,174 size 105x23; Text '工装电磁铁'
   TextField "文本域_5" at 410,226 size 105x23; Text '吸取电磁阀'
   TextField "文本域_7" at 408,278 size 145x23; Text '下压气缸电磁阀'
   TextField "文本域_8" at 410,381 size 38x23; Text 'FFU'
   TextField "文本域_9" at 410,434 size 45x23; Text '照明'
   Rectangle "矩形_3" at 234,113 size 101x35
      Appearance <- "备用_3(1)"
   Rectangle "矩形_4" at 234,166 size 101x35
      Appearance <- "工装电磁铁"
   Rectangle "矩形_5" at 234,219 size 101x35
      Appearance <- "吸取螺丝电磁阀"
   Rectangle "矩形_6" at 234,272 size 101x35
      Appearance <- "下压气缸电磁阀"
   Rectangle "矩形_7" at 234,378 size 101x35
      Appearance <- "FFU"
   Rectangle "矩形_8" at 234,429 size 101x35
      Appearance <- "照明"
   Rectangle "矩形_9" at 234,325 size 101x35
      Appearance <- "备用(9)"
   TextField "文本域_10" at 408,329 size 85x23; Text '电批测试'
   Button "按钮_1" at 622,323 size 100x40; TextOff '开启'
      on Press: SetBit("HMI_MU_HMI电批启动")
      on Release: ResetBit("HMI_MU_HMI电批启动")

screen "当前报警" 800x480, template "按钮_1"
   GraphicView "图形视图_2" at 159,185 size 50x50; Picture "图形_2"
   AlarmView "报警视图_1" at 218,63 size 572x410

screen "用户" 800x480, template "按钮"
   GraphicView "图形视图_2" at 156,308 size 50x50; Picture "图形_2"
   UserView "用户视图_1" at 220,67 size 577x409

screen "配方" 800x480, template "按钮"
   GraphicView "图形视图_2" at 153,244 size 50x50; Picture "图形_2"
   TextField "文本域_2" at 219,97 size 85x23; Text '产品选择'
   SymbolicIOField "符号 I/O 域_1" at 220,130 size 160x35; TextOn '1'; TextOff '0'; TextList "产品切换"
      ProcessValue <- "CAOZUO_Index"
   Button "HmiScreenItemData_1" at 395,130 size 127x35; TextOff '读取'; PictureOn "图形_13"; PictureOff "图形_38"
      on Release: ResetBit("CAOZUO_READ_REQ"); ActivateScreen("配方_1", 0)
      on Press: SetBit("CAOZUO_READ_REQ")

screen "配方_1" 800x480, template "按钮"
   GraphicView "图形视图_2" at 153,244 size 50x50; Picture "图形_2"
   TextField "文本域_2" at 219,97 size 85x23; Text '产品选择'
   SymbolicIOField "符号 I/O 域_1" at 220,130 size 160x35; TextOn '1'; TextOff '0'; TextList "产品切换"
      ProcessValue <- "CAOZUO_Index"
   IOField "I/O 域_5" at 220,222 size 160x35; FormatPattern ??????????
      ProcessValue <- "UDPT_加工文件名称"
   TextField "文本域_10" at 219,182 size 85x23; Text '产品名称'
   Button "HmiScreenItemData_2" at 395,222 size 127x35; TextOff '写入'; PictureOn "图形_13"; PictureOff "图形_38"
      on Release: ResetBit("CAOZUO_WRITE_REQ")
      on Press: SetBit("CAOZUO_WRITE_REQ")
   IOField "I/O 域_1" at 220,317 size 160x35; FormatPattern s99
      ProcessValue <- "UDPT_加工螺丝数量"
   TextField "文本域_1" at 220,284 size 105x23; Text '锁螺丝个数'

Template "按钮_1" 800x480
   Group "Group" at 0,0 size 799x59; Picture "LOGO"
   GraphicView "模板_图形视图_2" at 0,0 size 200x59; Picture "复赛"
   Button "HmiScreenItemData_1" at 11,68 size 143x47; TextOn '上一页'; TextOff '上一页'; PictureOff "图形_16"; PictureOn "图形_16"
      on Release: ActivateScreen("主页", 0)
   Button "HmiScreenItemData_5" at 11,127 size 143x47; TextOn '信号监控'; TextOff '补螺丝功能'; PictureOn "Navigates to SIMATIC PLC 监视表 for TP700 Comfort 14.0.1.0"; PictureOff "Navigates to SIMATIC PLC 监视表 for TP700 Comfort 14.0.1.0"; Authorization "User"
      on Release: ActivateScreen("补螺丝功能", 0)
   Button "HmiScreenItemData_11" at 11,247 size 143x47; TextOn '历史报警'; TextOff '历史报警'; PictureOn "Navigates to 项目信息 for TP700 Comfort 14.0.1.0"; PictureOff "Navigates to 项目信息 for TP700 Comfort 14.0.1.0"
      on Release: ActivateScreen("报警历史", 0)
   Button "HmiScreenItemData_7" at 11,188 size 143x47; TextOn '当前报警'; TextOff '当前报警'; PictureOn "Navigates to 系统信息 for TP700 Comfort 14.0.1.0"; PictureOff "Navigates to 系统信息 for TP700 Comfort 14.0.1.0"
      on Release: ActivateScreen("当前报警", 0)
   Button "HmiScreenItemData_4" at 11,311 size 143x47; TextOff '用户管理'; Authorization "User"; PictureOff "Navigates to 用户管理 for TP700 Comfort 14.0.1.0"; PictureOn "Navigates to 用户管理 for TP700 Comfort 14.0.1.0"
      on Release: ActivateScreen("用户", 0)
   Button "HmiScreenItemData_2" at 12,373 size 143x47; TextOff '系统设置'; PictureOff "图形_18"; PictureOn "图形_18"
      on Release: ActivateScreen("系统设置", 0)
   IOField "模板_I/O 域_1" at 258,13 size 85x32; FormatPattern ????????????????????????????????????????????????????????????????????????????????
      ProcessValue <- "HMI_MU_PLC 配方名称"
   IOField "模板_I/O 域_2" at 362,15 size 35x30; FormatPattern 99
      ProcessValue <- "HMI_MU_PLC 程序号"
   TextField "文本域_6" at 410,16 size 91x29; Text '回原位中'
      Visibility <- "回原位中"
   TextField "文本域_2" at 501,16 size 91x29; Text '请回原位'
      Visibility <- "回原位标志位"
      Appearance <- "回原位标志位"
   TextField "文本域_1" at 410,16 size 111x29; Text '回原位完成'
      Visibility <- "回原位标志位"
   DateTimeField "模板_日期/时间域_1" at 597,20 size 201x21
   GraphicView "模板_图形视图_1" at 0,0 size 102x59; Picture "33"
   GraphicView "模板_图形视图_3" at 102,0 size 697x59; Picture "33"

